   Button "Button_70" at 788,457 size 126x262; TextOff 'Text'
      on Release: function_efd93a16("Tank 2S Status", 168, 315, -1, 0, 1)
      Appearance <- "504_Tank Grouping_DB2020_RUN TANK 5"
   Button "Button_66" at 921,457 size 126x261; TextOff 'Text'
      on Release: function_efd93a16("Tank 1S Status", 168, 315, -1, 0, 1)
      Appearance <- "504_Tank Grouping_DB2020_RUN TANK 3"
   Button "Button_61" at 1093,328 size 130x248; TextOff 'Text'
      on Release: function_efd93a16("Tank FP Status", 168, 315, -1, 0, 1)
      Appearance <- "504_Tank Grouping_DB2020_RUN TANK 1"
   Button "Button_62" at 919,205 size 126x242; TextOff 'Text'
      on Release: function_efd93a16("Tank 1P Status", 168, 315, -1, 0, 1)
      Appearance <- "504_Tank Grouping_DB2020_RUN TANK 2"
   Button "Button_68" at 789,202 size 126x246; TextOff 'Text'
      on Release: function_efd93a16("Tank 2P Status", 168, 315, -1, 0, 1)
      Appearance <- "504_Tank Grouping_DB2020_RUN TANK 4"
   Button "Button_72" at 654,205 size 126x242; TextOff 'Text'
      on Release: function_efd93a16("Tank 3P Status", 168, 315, -1, 0, 1)
      Appearance <- "504_Tank Grouping_DB2020_RUN TANK 6"
   Button "Button_76" at 524,205 size 126x243; TextOff 'Text'
      on Release: function_efd93a16("Tank 4P Status", 168, 315, -1, 0, 1)
      Appearance <- "504_Tank Grouping_DB2020_RUN TANK 8"
   Button "Button_78" at 392,206 size 126x241; TextOff 'Text'
      on Release: function_efd93a16("Tank 5P Status", 168, 315, -1, 0, 1)
      Appearance <- "504_Tank Grouping_DB2020_RUN TANK 10"
   Button "Button_84" at 259,204 size 126x244; TextOff 'Text'
      on Release: function_efd93a16("Tank 6P Status", 168, 315, -1, 0, 1)
      Appearance <- "504_Tank Grouping_DB2020_RUN TANK 12"
   Group "Group_1" at 711,46 size 50x27; FormatPattern 999; Unit h
   Group "Group_2" at 605,46 size 57x27; FormatPattern 999; Unit h
   Button "HmiScreenItemData_5" at 180,144 size 116x50; TextOn 'Back'; TextOff 'Tank Status'
      on Release: function_efd93a16("Tank Status", 400, 250, -1, -1, 1)
   Button "Button_10" at 14,93 size 153x55; TextOff 'Text'
      on Release: function_efd93a16("Salinity - Acceptance", 168, 315, -1, 0, 1)
      Visibility <- "2068_Sys_Status_Data_SAL_VALID"
   Button "Button_12" at 14,93 size 153x54; TextOff 'Text'
      on Release: function_efd93a16("Tank Times", 300, 200, -1, 0, 1)
      Visibility <- "2068_Sys_Status_Data_Times Visibil"
   IOField "I/O field_29" at 664,46 size 45x27; FormatPattern 99; Unit h
      Visibility <- "2110_BTCS_CNTRL_DB_BTCS_STATE"
      ProcessValue <- "Sequence Times_DB_Treatment Timer_Hours Left"
   IOField "I/O field_30" at 664,46 size 45x27; FormatPattern 99; Unit h
      Visibility <- "2110_BTCS_CNTRL_DB_BTCS_STATE"
      ProcessValue <- "Sequence Times_DB_Pre-Dwell Timer_Hours Left"
   Button "Button_59" at 298,44 size 240x30; TextOn 'TB3 Enabled'; TextOff 'BWT System Shutting Down'
      Visibility <- "2110_BTCS_CNTRL_DB_BTCS_STATE"
   Button "Button_60" at 299,44 size 240x30; TextOn 'TB3 Enabled'; TextOff 'BWT System Enabled'
      Visibility <- "2110_BTCS_CNTRL_DB_BTCS_STATE"
   IOField "I/O field_15" at 711,46 size 50x27; FormatPattern 99; Unit m
      Visibility <- "2110_BTCS_CNTRL_DB_BTCS_STATE"
      ProcessValue <- "Sequence Times_DB_Treatment Timer_Minutes Left"
   IOField "I/O field_16" at 711,46 size 50x27; FormatPattern 99; Unit m
      Visibility <- "2110_BTCS_CNTRL_DB_BTCS_STATE"
      ProcessValue <- "Sequence Times_DB_Pre-Dwell Timer_Minutes Left"
   IOField "I/O field_17" at 605,46 size 57x27; FormatPattern 999; Unit d
      Visibility <- "2110_BTCS_CNTRL_DB_BTCS_STATE"
      ProcessValue <- "Sequence Times_DB_Treatment Timer_Days Left"
   IOField "I/O field_18" at 605,46 size 57x27; FormatPattern 999; Unit d
      Visibility <- "2110_BTCS_CNTRL_DB_BTCS_STATE"
      ProcessValue <- "Sequence Times_DB_Pre-Dwell Timer_Days Left"

screen "Balast Water Treatment Setup" 1280x800, template "Template"
   Button "HmiScreenItemData_1" at 1,1 size 150x40; TextOn 'Back'; TextOff 'Main Index'
      on Release: ActivateScreen("02 Main Index", 0)
   Button "HmiScreenItemData_8" at 276,83 size 219x27; TextOn 'Back'; TextOff 'Plant Operation'
   Button "HmiScreenItemData_23" at 282,116 size 150x47; TextOn 'Back'; TextOff 'Accept & Launch'; Authorization "Operate"
      Appearance <- "2110_BTCS_CNTRL_DB_BTCS_STATE"
      on Release: function_efd93a16("BWTS Start Confirm", 400, 200, -1, -1, 1)
      ObjectEnable <- "82_To_HMI_CRNT_MODE_GCU"
   Button "HmiScreenItemData_14" at 828,54 size 416x27; TextOn 'Back'; TextOff 'Treatment Durations'
   TextField "Text field_1" at 925,535 size 220x18; Text 'Tank Water Low Level (LT421)'
   TextField "Text field_2" at 925,573 size 220x18; Text 'Tank Water Low Level (LT422)'
   TextField "Text field_3" at 925,501 size 85x18; Text 'Description'
   TextField "Text field_5" at 925,611 size 215x18; Text 'De-Oxygenation DO Set Point'
   TextField "Text field_6" at 1164,501 size 67x18; Text 'Setpoint'
   Button "HmiScreenItemData_15" at 915,461 size 329x27; TextOn 'Back'; TextOff 'Ballast Tank Treatment Settings'
   IOField "I/O field_4" at 1153,530 size 80x28; Authorization "Operate"; FormatPattern 999.9; Unit  %
      ProcessValue <- "2084_Setpoints_LT421_Lo"
   IOField "I/O field_5" at 1153,568 size 80x28; Authorization "Operate"; FormatPattern 999.9; Unit  %
      ProcessValue <- "2084_Setpoints_LT422_Lo"
   IOField "I/O field_6" at 1153,606 size 80x28; Authorization "Operate"; FormatPattern 99.9; Unit  mg/l
      ProcessValue <- "2084_Setpoints_DO_SP"
   Button "HmiScreenItemData_16" at 482,461 size 334x27; TextOn 'Back'; TextOff 'Manual Ballast Tank Selection'
   Button "HmiScreenItemData_34" at 43,83 size 230x27; TextOn 'Back'; TextOff 'Plant Mode of Operation'
   Button "HmiScreenItemData_18" at 43,54 size 452x27; TextOn 'Back'; TextOff 'Ballast Water Treatment'
   Button "HmiScreenItemData_40" at 508,54 size 300x27; TextOn 'Back'; TextOff 'Treatment Status'
   TextField "Text field_14" at 837,94 size 85x18; Text 'Description'
   TextField "Text field_17" at 1054,94 size 67x18; Text 'Setpoint'
   IOField "I/O field_10" at 1040,132 size 92x27; Authorization "Operating Mode"; FormatPattern 999.99; Unit  Days
      ProcessValue <- "2115_VOYAGE_TIME_DAYS_VOYAGE_DAYS"
   IOField "I/O field_12" at 1040,267 size 79x28; Authorization "Commissioning"; FormatPattern 999; Unit  Hrs
      ProcessValue <- "2110_BTCS_CNTRL_DB_DE_OX_HRS"
   IOField "I/O field_13" at 1040,335 size 79x28; Authorization "Commissioning"; FormatPattern 999; Unit  Hrs
      ProcessValue <- "2110_BTCS_CNTRL_DB_DWELL_HRS"
   IOField "I/O field_14" at 1040,369 size 79x28; Authorization "Commissioning"; FormatPattern 999; Unit  Hrs
      ProcessValue <- "2110_BTCS_CNTRL_DB_RE_OX_HRS"
   IOField "I/O field_15" at 1040,403 size 79x28; Authorization "Commissioning"; FormatPattern 999; Unit  Hrs
      ProcessValue <- "2110_BTCS_CNTRL_DB_POST_DWELL_HRS"
   Button "HmiScreenItemData_11" at 836,128 size 203x35; TextOn 'Back'; TextOff 'Voyage A'
   Button "HmiScreenItemData_12" at 836,233 size 203x28; TextOn 'Back'; TextOff 'Pre Dwell Time'
   Button "HmiScreenItemData_13" at 836,267 size 203x28; TextOn 'Back'; TextOff 'De-Oxygenation Minimum Time'
   Button "HmiScreenItemData_43" at 836,335 size 203x28; TextOn 'Back'; TextOff 'Dwell Time'
   Button "HmiScreenItemData_44" at 836,369 size 203x28; TextOn 'Back'; TextOff 'Re-Oxygenation Time'
   Button "HmiScreenItemData_45" at 836,403 size 203x28; TextOn 'Back'; TextOff 'Post Dwell Time'
   IOField "I/O field_17" at 1060,169 size 79x28; Authorization "User administration"; FormatPattern 999; Unit  Hrs
      ProcessValue <- "2110_BTCS_CNTRL_DB_TOT_SEQ_HRS"
   Button "HmiScreenItemData_42" at 836,169 size 203x28; TextOn 'Back'; TextOff 'Total Treatment Time'
   Button "HmiScreenItemData_47" at 482,461 size 418x27; TextOn 'Back'; TextOff 'Automatic Ballast Tank Selection'
   Button "HmiScreenItemData_9" at 525,88 size 220x30; TextOn 'Back'; TextOff 'Pre Dwell Time Completed'
   Button "HmiScreenItemData_17" at 525,148 size 220x30; TextOn 'Back'; TextOff 'De-Oxygenation Completed'
   Button "HmiScreenItemData_38" at 525,178 size 220x30; TextOn 'Back'; TextOff 'Dwell Time Completed'
   Button "HmiScreenItemData_39" at 525,238 size 220x30; TextOn 'Back'; TextOff 'Re-Oxygenation Completed'
   Button "HmiScreenItemData_41" at 525,269 size 220x30; TextOn 'Back'; TextOff 'Post Dwell Time Completed'
   Button "HmiScreenItemData_46" at 525,118 size 220x30; TextOn 'Back'; TextOff 'Inert Gas Transfer Active'
   Button "HmiScreenItemData_48" at 525,208 size 220x30; TextOn 'Back'; TextOff 'Ambient Air Transfer Active'
   Button "HmiScreenItemData_52" at 525,118 size 220x30; TextOn 'Back'; TextOff 'IG Transfer Completed'
   Button "HmiScreenItemData_53" at 525,208 size 220x30; TextOn 'Back'; TextOff 'Ambient Air Transfer Completed'
   Button "HmiScreenItemData_3" at 1129,1 size 150x40; TextOn 'I&A Compressor Ok'; TextOff 'Back'
      on Release: function_efd93a16()
   TextField "Text field_11" at 1179,94 size 36x18; Text 'ETA'
   IOField "I/O field_16" at 1156,233 size 83x28; Authorization "User administration"; FormatPattern 999; Unit  min
      ProcessValue <- "2102_TIME_CALCS_DB_PRE_DWELL_MINS_RMNG"
   IOField "I/O field_18" at 1156,267 size 83x28; Authorization "User administration"; FormatPattern 999; Unit  min
   IOField "I/O field_19" at 1156,335 size 83x28; FormatPattern 999; Unit  min
      ProcessValue <- "2102_TIME_CALCS_DB_DWELL_MINS_RMNG"
   IOField "I/O field_20" at 1156,369 size 83x28; FormatPattern 999; Unit  min
      ProcessValue <- "2102_TIME_CALCS_DB_RE_OX_MINS_RMNG"
   IOField "I/O field_21" at 1156,403 size 83x28; FormatPattern 999; Unit  min
      ProcessValue <- "2102_TIME_CALCS_DB_POST_DWELL_MINS_RMNG"
   IOField "I/O field_22" at 1156,169 size 83x28; Authorization "User administration"; FormatPattern 999; Unit  Hrs
      ProcessValue <- "2110_BTCS_CNTRL_DB_RMNG_SEQ_HRS"
   Rectangle "Rectangle_25" at 281,165 size 179x59
      Visibility <- "2100_AUTO_SEQ_DB_SEQ_RNG"
   Button "HmiScreenItemData_4" at 282,172 size 150x47; TextOn 'Back'; TextOff 'Abort & Stop'; Authorization "Operate"
      Appearance <- "2110_BTCS_CNTRL_DB_BTCS_STATE"
      on Release: function_efd93a16("BWTS Stop Confirm", 400, 200, -1, -1, 1)
      ObjectEnable <- "82_To_HMI_CRNT_MODE_GCU"
   Circle "Circle_9" at 453,125 size 29x29
      Appearance <- "2110_BTCS_CNTRL_DB_BTCS_STATE"
   Circle "Circle_1" at 453,181 size 29x29
      Appearance <- "2110_BTCS_CNTRL_DB_BTCS_STATE"
   TextField "Text field_60" at 936,698 size 290x35; Text 'SALINITY ACCEPTED'
      Visibility <- "2068_Sys_Status_Data_SAL_VALID"
   Circle "Circle_19" at 220,233 size 29x29
      Appearance <- "150_GCU_LCL_CNTRL_DB_LCL_CNTRL_ACTV"
   Circle "Circle_20" at 220,180 size 29x29
      Appearance <- "82_To_HMI_CRNT_MODE_GCU"
   Button "HmiScreenItemData_36" at 49,170 size 150x51; TextOn 'Back'; TextOff 'Manual'; Authorization "Operate"
      on Press: function_b14e0dd5("80_From_HMI_Request_Manual", 0); ResetBit("150_GCU_LCL_CNTRL_DB_LCL_CNTRL_ACTV")
   Circle "Circle_21" at 220,126 size 29x29
      Appearance <- "82_To_HMI_CRNT_MODE_GCU"
   Button "HmiScreenItemData_37" at 49,116 size 150x51; TextOn 'Back'; TextOff 'Full Auto'; Authorization "Operate"
      on Press: function_b14e0dd5("80_From_HMI_Request_Auto", 0); ResetBit("150_GCU_LCL_CNTRL_DB_LCL_CNTRL_ACTV")
   Button "HmiScreenItemData_49" at 49,225 size 150x51; TextOn 'Back'; TextOff 'Local Auto'; Authorization "User administration"
      on Press: InvertBit("150_GCU_LCL_CNTRL_DB_LCL_CNTRL_ACTV"); function_b14e0dd5("80_From_HMI_Request_Auto", 0); ResetBit("80_From_HMI_Request_Manual")
   Circle "Circle_22" at 220,126 size 29x29
      Visibility <- "150_GCU_LCL_CNTRL_DB_LCL_CNTRL_ACTV"
   Circle "Circle_30" at 220,233 size 29x29
      Visibility <- "82_To_HMI_CRNT_MODE_GCU"
   Button "Button_4" at 493,507 size 100x23; TextOff 'FPT'; Authorization "Operate"
      on Press: function_b14e0dd5("504_Tank Grouping_DB2020_TANK ACTIV 1", 0)
      Appearance <- "504_Tank Grouping_DB2020_TANK ACTIV 1"
   Button "HmiScreenItemData_50" at 1156,297 size 83x35; TextOn 'Back'; TextOff 'Boost'; Authorization "Commissioning"
      on Press: InvertBit("Sequence Times_DB_Boost")
      Visibility <- "user_group"
      Appearance <- "Sequence Times_DB_Boost"
   IOField "I/O field_1" at 1040,301 size 79x28; Authorization "Commissioning"; FormatPattern 999; Unit  Hrs
      ProcessValue <- "2110_BTCS_CNTRL_DB_DE_OX_SP_HRS"
   Button "HmiScreenItemData_6" at 836,301 size 203x28; TextOn 'Back'; TextOff 'De-Oxygenation Setpoint Time'
   Rectangle "Rectangle_21" at 917,659 size 327x40
      Appearance <- "2068_Sys_Status_Data_SAL_VALID"
   TextField "Text field_48" at 916,664 size 128x30; Text 'Salinity Value:'
   IOField "I/O field_31" at 1036,664 size 74x30; FormatPattern 99.9; Unit psu
      ProcessValue <- "80_From_HMI_SAL_VALUE"
   Button "HmiScreenItemData_35" at 1108,664 size 135x30; TextOn 'Back'; TextOff 'Confirm Salinity'
      on Release: function_efd93a16("Salinity - Acceptance", 0, 0, 1, 3, 1)
   Group "Group_18" at 921,659 size 322x40
   Group "Group" at 916,659 size 327x40; Authorization "Operate"
   Button "HmiScreenItemData_7" at 1156,85 size 83x35; TextOn 'CONTINUE'; TextOff 'Continue'; Authorization "Operating Mode"
      on Press: InvertBit("80_From_HMI_TIMER RST Supres")
      Appearance <- "80_From_HMI_TIMER RST Supres"
   IOField "I/O field_25" at 1040,201 size 79x28; Authorization "User administration"; FormatPattern 999.9; Unit  Hrs
      ProcessValue <- "504_Tank Grouping_DB2020_Sequence Time m Offset_Real"
   Button "HmiScreenItemData_2" at 836,201 size 203x28; TextOn 'Back'; TextOff 'Differential Treatment Time'
   IOField "I/O field_3" at 1156,201 size 83x28; Authorization "User administration"; FormatPattern 999; Unit  min
      ProcessValue <- "504_Tank Grouping_DB2020_Diff Time Remain"
   Button "Button_1" at 817,594 size 79x32; TextOff '3'; Authorization "Operate"
      on Press: function_b14e0dd5("504_Tank Grouping_DB2020_GROUP ACTIV 3", 0)
      Appearance <- "504_Tank Grouping_DB2020_GROUP ACTIVE INT 3"
   Button "Button_2" at 817,628 size 79x32; TextOff '4'; Authorization "Operate"
      on Press: function_b14e0dd5("504_Tank Grouping_DB2020_GROUP ACTIV 4", 0)
      Appearance <- "504_Tank Grouping_DB2020_GROUP ACTIVE INT 4"
   Button "Button_10" at 818,662 size 79x32; TextOff '5'; Authorization "Operate"
      on Press: function_b14e0dd5("504_Tank Grouping_DB2020_GROUP ACTIV 5", 0)
      Appearance <- "504_Tank Grouping_DB2020_GROUP ACTIVE INT 5"
   Button "Button_11" at 818,696 size 79x32; TextOff '6'; Authorization "Operate"
      on Press: function_b14e0dd5("504_Tank Grouping_DB2020_GROUP ACTIV 6", 0)
      Appearance <- "504_Tank Grouping_DB2020_GROUP ACTIVE INT 6"
   Button "Button_12" at 818,731 size 79x32; TextOff '7'; Authorization "Operate"
      on Press: function_b14e0dd5("504_Tank Grouping_DB2020_GROUP ACTIV 7", 0)
      Appearance <- "504_Tank Grouping_DB2020_GROUP ACTIVE INT 7"
   IOField "I/O field_37" at 183,323 size 90x29; Authorization "Commissioning"; FormatPattern 999; Unit  step
      ProcessValue <- "2110_BTCS_CNTRL_DB_BTCS_STEP"
   Button "HmiScreenItemData_10" at 43,323 size 137x29; TextOn 'Back'; TextOff 'BWTS Step'
   Button "HmiScreenItemData_51" at 43,358 size 137x29; TextOn 'Back'; TextOff 'BWTS State'
   Button "HmiScreenItemData_54" at 276,323 size 532x29; TextOn 'Back'; TextOff 'IGG STEP'; TextList "STEP LIST BTCS"
      ProcessValue <- "2110_BTCS_CNTRL_DB_BTCS_STEP"
   Button "HmiScreenItemData_55" at 276,358 size 532x29; TextOn 'Back'; TextOff 'IGG STEP'; TextList "STATE LIST BTCS"
      ProcessValue <- "2110_BTCS_CNTRL_DB_BTCS_STATE"
   Circle "Circle_2" at 421,496 size 26x26
      Appearance <- "80_From_HMI_BWT_BYPASS"
   Button "HmiScreenItemData_57" at 88,494 size 304x33; TextOn 'Back'; TextOff 'Ballast Water Treatment'; Authorization "Operate"
      on Press: InvertBit("80_From_HMI_BWT_BYPASS(1)"); ResetBit("80_From_HMI_CRG_BLNK_MODE(1)")
      Appearance <- "80_From_HMI_BWT_BYPASS(1)"
      ObjectEnable <- "100_GCU_AUTO_SEQ_DB_CRNT_STEP"
   Circle "Circle_3" at 421,534 size 26x26
      Appearance <- "80_From_HMI_CRG_BLNK_MODE"
   Button "HmiScreenItemData_58" at 88,532 size 304x33; TextOn 'Back'; TextOff 'Cargo Blanketing'; Authorization "Operate"
      on Press: InvertBit("80_From_HMI_CRG_BLNK_MODE(1)"); ResetBit("80_From_HMI_BWT_BYPASS(1)")
      Appearance <- "80_From_HMI_CRG_BLNK_MODE(1)"
      ObjectEnable <- "100_GCU_AUTO_SEQ_DB_CRNT_STEP"
   Button "HmiScreenItemData_56" at 41,461 size 425x27; TextOn 'Back'; TextOff 'Inert Gas Transfer Mode'
   Button "Button_7" at 817,526 size 79x32; TextOff '1'; Authorization "Operate"
      on Press: function_b14e0dd5("504_Tank Grouping_DB2020_GROUP ACTIV 1", 0)
      Appearance <- "504_Tank Grouping_DB2020_GROUP ACTIVE INT 1"
   Button "Button_8" at 817,560 size 79x32; TextOff '2'; Authorization "Operate"
      on Press: function_b14e0dd5("504_Tank Grouping_DB2020_GROUP ACTIV 2", 0)
      Appearance <- "504_Tank Grouping_DB2020_GROUP ACTIVE INT 2"
   Button "Button_9" at 493,539 size 100x23; TextOff 'TANK - 1P'; Authorization "Operate"
      on Press: function_b14e0dd5("504_Tank Grouping_DB2020_TANK ACTIV 2", 0)
      Appearance <- "504_Tank Grouping_DB2020_TANK ACTIV 2"
   Button "Button_14" at 493,571 size 100x23; TextOff 'TANK - 2P'; Authorization "Operate"
      on Press: function_b14e0dd5("504_Tank Grouping_DB2020_TANK ACTIV 4", 0)
      Appearance <- "504_Tank Grouping_DB2020_TANK ACTIV 4"
   Button "Button_15" at 493,603 size 100x23; TextOff 'TANK - 3P'; Authorization "Operate"
      on Press: function_b14e0dd5("504_Tank Grouping_DB2020_TANK ACTIV 6", 0)
      Appearance <- "504_Tank Grouping_DB2020_TANK ACTIV 6"
   Button "Button_16" at 493,636 size 100x23; TextOff 'TANK - 4P'; Authorization "Operate"
      on Press: function_b14e0dd5("504_Tank Grouping_DB2020_TANK ACTIV 8", 0)
      Appearance <- "504_Tank Grouping_DB2020_TANK ACTIV 8"
   Button "Button_17" at 493,668 size 100x23; TextOff 'TANK - 5P'; Authorization "Operate"
      on Press: function_b14e0dd5("504_Tank Grouping_DB2020_TANK ACTIV 10", 0)
      Appearance <- "504_Tank Grouping_DB2020_TANK ACTIV 10"
   Button "Button_18" at 493,700 size 100x23; TextOff 'TANK - 6P'; Authorization "Operate"
      on Press: function_b14e0dd5("504_Tank Grouping_DB2020_TANK ACTIV 12", 0)
      Appearance <- "504_Tank Grouping_DB2020_TANK ACTIV 12"
   Button "Button_19" at 493,733 size 100x23; TextOff 'TANK - APT'; Authorization "Operate"
      on Press: function_b14e0dd5("504_Tank Grouping_DB2020_TANK ACTIV 14", 0)
      Appearance <- "504_Tank Grouping_DB2020_TANK ACTIV 14"
   Button "Button_20" at 706,539 size 100x23; TextOff 'TANK - 1S'; Authorization "Operate"
      on Press: function_b14e0dd5("504_Tank Grouping_DB2020_TANK ACTIV 3", 0)
      Appearance <- "504_Tank Grouping_DB2020_TANK ACTIV 3"
   Button "Button_21" at 706,571 size 100x23; TextOff 'TANK - 2S'; Authorization "Operate"
      on Press: function_b14e0dd5("504_Tank Grouping_DB2020_TANK ACTIV 5", 0)
      Appearance <- "504_Tank Grouping_DB2020_TANK ACTIV 5"
   Button "Button_22" at 706,603 size 100x23; TextOff 'TANK - 3S'; Authorization "Operate"
      on Press: function_b14e0dd5("504_Tank Grouping_DB2020_TANK ACTIV 7", 0)
      Appearance <- "504_Tank Grouping_DB2020_TANK ACTIV 7"
   Button "Button_23" at 706,635 size 100x23; TextOff 'TANK - 4S'; Authorization "Operate"
      on Press: function_b14e0dd5("504_Tank Grouping_DB2020_TANK ACTIV 9", 0)
      Appearance <- "504_Tank Grouping_DB2020_TANK ACTIV 9"
   Button "Button_24" at 706,667 size 100x23; TextOff 'TANK - 5S'; Authorization "Operate"
      on Press: function_b14e0dd5("504_Tank Grouping_DB2020_TANK ACTIV 11", 0)
      Appearance <- "504_Tank Grouping_DB2020_TANK ACTIV 11"
   Button "Button_25" at 706,700 size 100x23; TextOff 'TANK - 6S'; Authorization "Operate"
      on Press: function_b14e0dd5("504_Tank Grouping_DB2020_TANK ACTIV 13", 0)
      Appearance <- "504_Tank Grouping_DB2020_TANK ACTIV 13"
   IOField "I/O field_38" at 183,358 size 90x29; Authorization "Commissioning"; FormatPattern 9; Unit  state
      ProcessValue <- "2110_BTCS_CNTRL_DB_BTCS_STATE"
   Switch "Switch_8" at 776,732 size 32x29; CaptionText 'Switch'; TextOn 'ON'; TextOff 'OFF'; Authorization "User administration"; PictureOff "Design_5_PilotLight_Green_Off"; PictureOn "Design_5_PilotLight_Green_On"
      on Change: InvertBit("80_From_HMI_Test Tank Request")
      ProcessValue <- "504_Tank Grouping_DB2020_RUN"
      Visibility <- "user_group"
   Circle "Circle_31" at 621,507 size 20x20
      Visibility <- "504_Tank Grouping_DB2020_RUN TANK 1"
      Appearance <- "504_Tank Grouping_DB2020_RUN TANK 1"
   Circle "Circle_4" at 600,573 size 20x20
      Appearance <- "504_Tank Grouping_DB2020_GROUP of TANK 4"
   Circle "Circle_6" at 599,604 size 20x20
      Appearance <- "504_Tank Grouping_DB2020_GROUP of TANK 6"
   Circle "Circle_7" at 599,541 size 20x20
      Appearance <- "504_Tank Grouping_DB2020_GROUP of TANK 2"
   Circle "Circle_8" at 599,669 size 20x20
      Appearance <- "504_Tank Grouping_DB2020_GROUP of TANK 10"
   Circle "Circle_10" at 599,637 size 20x20
      Appearance <- "504_Tank Grouping_DB2020_GROUP of TANK 8"
   Circle "Circle_11" at 599,734 size 20x20
      Appearance <- "504_Tank Grouping_DB2020_GROUP of TANK 14"
   Circle "Circle_12" at 599,701 size 20x20
      Appearance <- "504_Tank Grouping_DB2020_GROUP of TANK 12"
   IOField "I/O field_8" at 599,544 size 20x14; FormatPattern 99
      ProcessValue <- "504_Tank Grouping_DB2020_GROUP of TANK 2"
   IOField "I/O field_9" at 599,576 size 20x14; FormatPattern 99
      ProcessValue <- "504_Tank Grouping_DB2020_GROUP of TANK 4"
   IOField "I/O field_26" at 599,607 size 20x14; FormatPattern 99
      ProcessValue <- "504_Tank Grouping_DB2020_GROUP of TANK 6"
   IOField "I/O field_28" at 599,640 size 20x14; FormatPattern 99
      ProcessValue <- "504_Tank Grouping_DB2020_GROUP of TANK 8"
   IOField "I/O field_30" at 599,672 size 20x14; FormatPattern 99
      ProcessValue <- "504_Tank Grouping_DB2020_GROUP of TANK 10"
   IOField "I/O field_33" at 599,704 size 20x14; FormatPattern 99
      ProcessValue <- "504_Tank Grouping_DB2020_GROUP of TANK 12"
   IOField "I/O field_35" at 599,737 size 20x14; FormatPattern 99
      ProcessValue <- "504_Tank Grouping_DB2020_GROUP of TANK 14"
   Circle "Circle_13" at 678,573 size 20x20
      Appearance <- "504_Tank Grouping_DB2020_GROUP of TANK 5"
   Circle "Circle_14" at 678,603 size 20x20
      Appearance <- "504_Tank Grouping_DB2020_GROUP of TANK 7"
   Circle "Circle_15" at 678,541 size 20x20
      Appearance <- "504_Tank Grouping_DB2020_GROUP of TANK 3"
   Circle "Circle_16" at 678,668 size 20x20
      Appearance <- "504_Tank Grouping_DB2020_GROUP of TANK 11"
   Circle "Circle_17" at 678,636 size 20x20
      Appearance <- "504_Tank Grouping_DB2020_GROUP of TANK 9"
   Circle "Circle_18" at 678,701 size 20x20
      Appearance <- "504_Tank Grouping_DB2020_GROUP of TANK 13"
   IOField "I/O field_23" at 678,544 size 20x14; FormatPattern 99
      ProcessValue <- "504_Tank Grouping_DB2020_GROUP of TANK 3"
   IOField "I/O field_24" at 678,576 size 20x14; FormatPattern 99
      ProcessValue <- "504_Tank Grouping_DB2020_GROUP of TANK 5"
   IOField "I/O field_27" at 678,606 size 20x14; FormatPattern 99
      ProcessValue <- "504_Tank Grouping_DB2020_GROUP of TANK 7"
   IOField "I/O field_29" at 678,639 size 20x14; FormatPattern 99
      ProcessValue <- "504_Tank Grouping_DB2020_GROUP of TANK 9"
   IOField "I/O field_32" at 678,671 size 20x14; FormatPattern 99
      ProcessValue <- "504_Tank Grouping_DB2020_GROUP of TANK 11"
   IOField "I/O field_34" at 678,704 size 20x14; FormatPattern 99
      ProcessValue <- "504_Tank Grouping_DB2020_GROUP of TANK 13"
   Circle "Circle_32" at 621,540 size 20x20
      Visibility <- "504_Tank Grouping_DB2020_RUN TANK 2"
      Appearance <- "504_Tank Grouping_DB2020_RUN TANK 2"
   Circle "Circle_33" at 656,540 size 20x20
      Visibility <- "504_Tank Grouping_DB2020_RUN TANK 3"
      Appearance <- "504_Tank Grouping_DB2020_RUN TANK 3"
   Circle "Circle_34" at 621,572 size 20x20
      Visibility <- "504_Tank Grouping_DB2020_RUN TANK 4"
      Appearance <- "504_Tank Grouping_DB2020_RUN TANK 4"
   Circle "Circle_35" at 656,572 size 20x20
      Visibility <- "504_Tank Grouping_DB2020_RUN TANK 5"
      Appearance <- "504_Tank Grouping_DB2020_RUN TANK 5"
   Circle "Circle_36" at 621,604 size 20x20
      Visibility <- "504_Tank Grouping_DB2020_RUN TANK 6"
      Appearance <- "504_Tank Grouping_DB2020_RUN TANK 6"
   Circle "Circle_37" at 656,604 size 20x20
      Visibility <- "504_Tank Grouping_DB2020_RUN TANK 7"
      Appearance <- "504_Tank Grouping_DB2020_RUN TANK 7"
   Circle "Circle_38" at 621,636 size 20x20
      Visibility <- "504_Tank Grouping_DB2020_RUN TANK 8"
      Appearance <- "504_Tank Grouping_DB2020_RUN TANK 8"
   Circle "Circle_39" at 656,636 size 20x20
      Visibility <- "504_Tank Grouping_DB2020_RUN TANK 9"
      Appearance <- "504_Tank Grouping_DB2020_RUN TANK 9"
   Circle "Circle_40" at 621,668 size 20x20
      Visibility <- "504_Tank Grouping_DB2020_RUN TANK 10"
      Appearance <- "504_Tank Grouping_DB2020_RUN TANK 10"
   Circle "Circle_41" at 656,668 size 20x20
      Visibility <- "504_Tank Grouping_DB2020_RUN TANK 11"
      Appearance <- "504_Tank Grouping_DB2020_RUN TANK 11"
   Circle "Circle_42" at 621,701 size 20x20
      Visibility <- "504_Tank Grouping_DB2020_RUN TANK 12"
      Appearance <- "504_Tank Grouping_DB2020_RUN TANK 12"
   Circle "Circle_43" at 656,701 size 20x20
      Visibility <- "504_Tank Grouping_DB2020_RUN TANK 13"
      Appearance <- "504_Tank Grouping_DB2020_RUN TANK 13"
   Circle "Circle_44" at 621,733 size 20x20
      Visibility <- "504_Tank Grouping_DB2020_RUN TANK 14"
      Appearance <- "504_Tank Grouping_DB2020_RUN TANK 14"
   TextField "Text field_7" at 648,740 size 136x18; Text 'Test Tank Request'
      Visibility <- "user_group"
   Rectangle "Rectangle_6" at 816,488 size 82x37
      Visibility <- "504_Tank Grouping_DB2020_SetGroupSR"
   Button "Button_13" at 819,491 size 76x31; TextOff 'Set Group'; Authorization "Parameter Change"
      on Press: function_b14e0dd5("504_Tank Grouping_DB2020_SetGroup", 0)
      Appearance <- "504_Tank Grouping_DB2020_GROUP SET"
   Button "HmiScreenItemData_5" at 41,576 size 426x27; TextOn 'Back'; TextOff 'Automatic Gas to Tank Valves Cycling'
   Button "HmiScreenItemData_19" at 370,722 size 83x35; TextOn 'ENABLE'; TextOff 'Enable'; Authorization "Operate"
      on Press: InvertBit("504_Tank Grouping_DB2020_Valve Cycle_Enable")
      Appearance <- "504_Tank Grouping_DB2020_Valve Cycle_Enable"
   TextField "Text field_8" at 54,652 size 254x18; Text 'Gas to Tank Valves Cycle Frequency'
   TextField "Text field_9" at 54,690 size 233x18; Text 'Gas to Tank Valves Cycle Length'
   TextField "Text field_10" at 54,618 size 85x18; Text 'Description'
   TextField "Text field_12" at 311,618 size 67x18; Text 'Setpoint'
   IOField "I/O field_39" at 310,649 size 70x28; Authorization "Operate"; FormatPattern 999; Unit h
      ProcessValue <- "504_Tank Grouping_DB2020_Valve Cycle_Period"
   IOField "I/O field_40" at 310,685 size 70x28; Authorization "Operate"; FormatPattern 9999; Unit s
      ProcessValue <- "504_Tank Grouping_DB2020_Valve Cycle_Length"
   TextField "Text field_13" at 385,618 size 58x18; Text 'Elapsed'
   IOField "I/O field_41" at 384,649 size 70x28; Authorization "Operate"; FormatPattern 999; Unit h
      ProcessValue <- "504_Tank Grouping_DB2020_Cycle Period_ET"
   IOField "I/O field_42" at 384,685 size 70x28; Authorization "Operate"; FormatPattern 9999; Unit s
      ProcessValue <- "504_Tank Grouping_DB2020_Cycle Length_ET"
   IOField "I/O field_48" at 1172,169 size 33x28; Authorization "User administration"; FormatPattern 99; Unit h
      ProcessValue <- "Sequence Times_DB_Treatment Timer_Hours Left"
   IOField "I/O field_51" at 1140,169 size 33x28; Authorization "User administration"; FormatPattern 99; Unit d
      ProcessValue <- "Sequence Times_DB_Treatment Timer_Days Left"
   IOField "I/O field_52" at 1204,169 size 35x28; Authorization "User administration"; FormatPattern 99; Unit m
      ProcessValue <- "Sequence Times_DB_Treatment Timer_Minutes Left"
   IOField "I/O field_43" at 1156,201 size 83x28; Authorization "User administration"; FormatPattern 999; Unit  min
      ProcessValue <- "504_Tank Grouping_DB2020_Diff Time Remain"
      Visibility <- "AlwaysTRUE"
   IOField "I/O field_44" at 1204,233 size 35x28; Authorization "User administration"; FormatPattern 99; Unit m
      ProcessValue <- "Sequence Times_DB_Pre-Dwell Timer_Minutes Left"
   IOField "I/O field_45" at 1172,233 size 33x28; Authorization "User administration"; FormatPattern 99; Unit h
      ProcessValue <- "Sequence Times_DB_Pre-Dwell Timer_Hours Left"
   IOField "I/O field_46" at 1140,233 size 33x28; Authorization "User administration"; FormatPattern 99; Unit d
      ProcessValue <- "Sequence Times_DB_Pre-Dwell Timer_Days Left"
   IOField "I/O field_47" at 1040,132 size 92x28; Authorization "Operating Mode"; FormatPattern 999.9; Unit  Days
      ProcessValue <- "Sequence Times_DB_Jurney Time"
   IOField "I/O field_49" at 1072,169 size 33x28; Authorization "User administration"; FormatPattern 99; Unit h
      ProcessValue <- "Sequence Times_DB_Treatment Timer_Hours"
   IOField "I/O field_50" at 1040,169 size 33x28; Authorization "User administration"; FormatPattern 99; Unit d
      ProcessValue <- "Sequence Times_DB_Treatment Timer_Days"
   IOField "I/O field_53" at 1104,169 size 35x28; Authorization "User administration"; FormatPattern 99; Unit m
      ProcessValue <- "Sequence Times_DB_Treatment Timer_Minutes"
   IOField "I/O field_54" at 1172,132 size 33x28; Authorization "User administration"; FormatPattern 99; Unit h
      ProcessValue <- "Sequence Times_DB_Jurney Timer_Hours Left"
   IOField "I/O field_55" at 1133,132 size 40x28; Authorization "User administration"; FormatPattern 999; Unit d
      ProcessValue <- "Sequence Times_DB_Jurney Timer_Days Left"
   IOField "I/O field_56" at 1204,132 size 35x28; Authorization "User administration"; FormatPattern 99; Unit m
      ProcessValue <- "Sequence Times_DB_Jurney Timer_Minutes Left"
   IOField "I/O field_57" at 1040,233 size 79x28; Authorization "Commissioning"; FormatPattern 9999.9; Unit  Hrs
      ProcessValue <- "Sequence Times_DB_Pre-Dwell Time"
   IOField "I/O field_58" at 1040,267 size 79x28; Authorization "Commissioning"; FormatPattern 999.9; Unit  Hrs
      ProcessValue <- "Sequence Times_DB_De-Ox Time"
   IOField "I/O field_59" at 1204,267 size 35x28; Authorization "User administration"; FormatPattern 99; Unit m
      ProcessValue <- "Sequence Times_DB_De-Ox Timer_Minutes Left"
   IOField "I/O field_60" at 1172,267 size 33x28; Authorization "User administration"; FormatPattern 99; Unit h
      ProcessValue <- "Sequence Times_DB_De-Ox Timer_Hours Left"
   IOField "I/O field_61" at 1140,267 size 33x28; Authorization "User administration"; FormatPattern 99; Unit d
      ProcessValue <- "Sequence Times_DB_De-Ox Timer_Days Left"
   IOField "I/O field_62" at 1040,301 size 79x28; Authorization "Commissioning"; FormatPattern 999.9; Unit  Hrs
      ProcessValue <- "Sequence Times_DB_De-Ox SP Time"
   IOField "I/O field_63" at 1040,335 size 79x28; Authorization "Commissioning"; FormatPattern 999.9; Unit  Hrs
      ProcessValue <- "Sequence Times_DB_Dwell Time"
   IOField "I/O field_64" at 1204,335 size 35x28; Authorization "User administration"; FormatPattern 99; Unit m
      ProcessValue <- "Sequence Times_DB_Dwell Timer_Minutes Left"
   IOField "I/O field_65" at 1172,335 size 33x28; Authorization "User administration"; FormatPattern 99; Unit h
      ProcessValue <- "Sequence Times_DB_Dwell Timer_Hours Left"
   IOField "I/O field_66" at 1140,335 size 33x28; Authorization "User administration"; FormatPattern 99; Unit d
      ProcessValue <- "Sequence Times_DB_Dwell Timer_Days Left"
   IOField "I/O field_2" at 1040,369 size 79x28; Authorization "Commissioning"; FormatPattern 999.9; Unit  Hrs
      ProcessValue <- "Sequence Times_DB_Re-Ox Time"
   IOField "I/O field_67" at 1204,369 size 35x28; Authorization "User administration"; FormatPattern 99; Unit m
      ProcessValue <- "Sequence Times_DB_Re-Ox Timer_Minutes Left"
   IOField "I/O field_68" at 1172,369 size 33x28; Authorization "User administration"; FormatPattern 99; Unit h
      ProcessValue <- "Sequence Times_DB_Re-Ox Timer_Hours Left"
   IOField "I/O field_69" at 1140,369 size 33x28; Authorization "User administration"; FormatPattern 99; Unit d
      ProcessValue <- "Sequence Times_DB_Re-Ox Timer_Days Left"
   IOField "I/O field_70" at 1040,403 size 79x28; Authorization "Commissioning"; FormatPattern 999.9; Unit  Hrs
      ProcessValue <- "Sequence Times_DB_Post-Dwell Time"
   IOField "I/O field_71" at 1204,403 size 35x28; Authorization "User administration"; FormatPattern 99; Unit m
      ProcessValue <- "Sequence Times_DB_Post-Dwell Timer_Minutes Left"
   IOField "I/O field_72" at 1172,403 size 33x28; Authorization "User administration"; FormatPattern 99; Unit h
      ProcessValue <- "Sequence Times_DB_Post-Dwell Timer_Hours Left"
   IOField "I/O field_73" at 1140,403 size 33x28; Authorization "User administration"; FormatPattern 99; Unit d
      ProcessValue <- "Sequence Times_DB_Post-Dwell Timer_Days Left"
   TextField "Text field_15" at 621,419 size 156x18; Text 'Treatment Timer Test'
      Visibility <- "user_group"
   Switch "Switch_1" at 774,411 size 32x29; CaptionText 'Switch'; TextOn 'ON'; TextOff 'OFF'; Authorization "User administration"; PictureOff "Design_5_PilotLight_Green_Off"; PictureOn "Design_5_PilotLight_Green_On"
      on Change: InvertBit("80_From_HMI_Jurney Start Simulator")
      Visibility <- "user_group"
      ProcessValue <- "80_From_HMI_Jurney Start Simulator"
   Circle "Circle_5" at 599,507 size 20x20
      Appearance <- "504_Tank Grouping_DB2020_GROUP of TANK 1"
   IOField "I/O field_7" at 599,510 size 20x14; FormatPattern 99
      ProcessValue <- "504_Tank Grouping_DB2020_GROUP of TANK 1"
   TextField "Text field_16" at 72,422 size 76x18; Text 'HeartBeat'
      Visibility <- "user_group"
   TextField "Text field_18" at 201,422 size 107x18; Text 'PLC HeartBeat'
      Visibility <- "user_group"
   Circle "Circle_45" at 40,414 size 26x26
      Appearance <- "CCR HMI HEART BEAT"
      Visibility <- "user_group"
   Circle "Circle_46" at 166,414 size 26x26
      Appearance <- "IGG PLC HEART BEAT"
      Visibility <- "user_group"
   TextField "Text field_19" at 445,403 size 133x18; Text 'Log IGG Simulator'
      Visibility <- "user_group"
   Switch "Switch_2" at 568,393 size 32x29; CaptionText 'Switch'; TextOn 'ON'; TextOff 'OFF'; Authorization "User administration"; PictureOff "Design_5_PilotLight_Green_Off"; PictureOn "Design_5_PilotLight_Green_On"
      on Change: InvertBit("68_Sys_Status_Data_LOG IGG Simulator")
      Visibility <- "user_group"
      ProcessValue <- "68_Sys_Status_Data_LOG IGG Simulator"
   TextField "Text field_20" at 445,435 size 136x18; Text 'Log GCU Simulator'
      Visibility <- "user_group"
   Switch "Switch_3" at 568,425 size 32x29; CaptionText 'Switch'; TextOn 'ON'; TextOff 'OFF'; Authorization "User administration"; PictureOff "Design_5_PilotLight_Green_Off"; PictureOn "Design_5_PilotLight_Green_On"
      on Change: InvertBit("68_Sys_Status_Data_LOG GCU Simulator")
      Visibility <- "user_group"
      ProcessValue <- "68_Sys_Status_Data_LOG GCU Simulator"
   Button "Button_5" at 53,722 size 210x35; TextOff 'PGC Setpoint Protection'
      on Press: function_efd93a16("PGC Setpoint Protection", 400, 200, -1, -1, 1)
   Button "Button_26" at 281,116 size 208x107; TextOff 'Text'
      on Release: function_efd93a16("Salinity - Acceptance", 168, 315, -1, 0, 1)
      Visibility <- "2068_Sys_Status_Data_SAL_VALID"
   Button "Button_27" at 280,115 size 204x107; TextOff 'Text'
      on Release: function_efd93a16("Tank Times", 300, 200, -1, 0, 1)
      Visibility <- "2068_Sys_Status_Data_Times Visibil"
   Group "Group_1" at 909,732 size 329x37
   IOField "I/O field_11" at 1156,201 size 83x28; Authorization "User administration"; FormatPattern 999; Unit  Hrs
      ProcessValue <- "2110_BTCS_CNTRL_DB_RMNG_SEQ_HRS"
   IOField "I/O field_74" at 1172,201 size 33x28; Authorization "User administration"; FormatPattern 99; Unit h
      ProcessValue <- "Sequence Times_DB_Offset Timer_Hours Left"
   IOField "I/O field_75" at 1140,201 size 33x28; Authorization "User administration"; FormatPattern 99; Unit d
      ProcessValue <- "Sequence Times_DB_Offset Timer_Days Left"
   IOField "I/O field_76" at 1204,201 size 35x28; Authorization "User administration"; FormatPattern 99; Unit m
      ProcessValue <- "Sequence Times_DB_Offset Timer_Minutes Left"
   Circle "Circle_23" at 764,91 size 24x24
      Appearance <- "2110_BTCS_CNTRL_DB_BTCS_STEP"
   Circle "Circle_24" at 764,120 size 24x24
      Appearance <- "100_GCU_AUTO_SEQ_DB_CRNT_STEP"
   Circle "Circle_25" at 764,150 size 24x24
      Appearance <- "2110_BTCS_CNTRL_DB_BTCS_STEP"
   Circle "Circle_26" at 764,180 size 24x24
      Appearance <- "2110_BTCS_CNTRL_DB_BTCS_STEP"
   Circle "Circle_27" at 764,210 size 24x24
      Appearance <- "100_GCU_AUTO_SEQ_DB_CRNT_STEP"
   Circle "Circle_28" at 764,240 size 24x24
      Appearance <- "2110_BTCS_CNTRL_DB_BTCS_STEP"
   Circle "Circle_29" at 764,270 size 24x24
      Appearance <- "2110_BTCS_CNTRL_DB_BTCS_STEP"
   TextField "Text field_34" at 980,733 size 187x35; Text 'TIMES VALID'
      Visibility <- "2102_TIME_CALCS_DB_TIMES_VALID"
   TextField "Text field_4" at 909,732 size 329x37; Text 'TIMES INVALID'
      Visibility <- "2102_TIME_CALCS_DB_TIMES_VALID"
   Rectangle "Rectangle_27" at 921,659 size 322x40
      Visibility <- "2068_Sys_Status_Data_SAL_CNF_CHK"
   TextField "Text field_62" at 925,664 size 156x30; Text 'Confirm Salinity? :'
      Visibility <- "2068_Sys_Status_Data_SAL_CNF_CHK"
   Button "Button_6" at 1086,664 size 67x30; TextOff 'YES'
      on Press: function_b14e0dd5("80_From_HMI_LOW_SAL_ACPT", 0)
      Visibility <- "2068_Sys_Status_Data_SAL_CNF_CHK"
   Button "Button_3" at 1166,664 size 67x30; TextOff 'NO'
      on Press: function_b14e0dd5("80_From_HMI_LOW_SAL_RJCT", 0)
      Visibility <- "2068_Sys_Status_Data_SAL_CNF_CHK"
   Rectangle "Rectangle_28" at 916,659 size 327x40
      Visibility <- "2100_AUTO_SEQ_DB_SEQ_RNG"
      Appearance <- "2102_TIME_CALCS_DB_RE_OX_SP_TMR_DN"
   TextField "Text field_49" at 920,664 size 211x30; Text 'Salinity Value :'
      Visibility <- "2100_AUTO_SEQ_DB_SEQ_RNG"
   IOField "I/O field_36" at 1131,664 size 95x30; Authorization "Operate"; FormatPattern 99.9; Unit psu
      ProcessValue <- "80_From_HMI_SAL_VALUE"
      Visibility <- "2100_AUTO_SEQ_DB_SEQ_RNG"

PopupScreen "Tank 1P Status" 885x425
   TrendView "Trend view_1" at 280,8 size 600x360
   TextField "Text field_4" at 20,136 size 86x22; Text 'Pressure:'
   IOField "I/O field_1" at 175,131 size 90x25; FormatPattern s999.9; Unit  mBar
      ProcessValue <- "20_TANKS_IP_DATA_RIO_01_FIRST_TANK_TANKS_PRESS"
   TextField "Text field_5" at 20,170 size 113x22; Text 'Water Level:'
   IOField "I/O field_2" at 175,165 size 90x25; FormatPattern 999.9; Unit  %
      ProcessValue <- "20_TANKS_IP_DATA_RIO_01_SECOND_TANK_BWT_LEVEL"
   TextField "Text field_6" at 20,204 size 137x22; Text 'MBG Flow Rate:'
   IOField "I/O field_3" at 175,199 size 90x25; FormatPattern 999.9; Unit  m³/hr
      ProcessValue <- "20_TANKS_IP_DATA_RIO_01_SECOND_TANK_MBG_FLOW"
   TextField "Text field_7" at 20,238 size 135x22; Text 'USD Flow Rate:'
   IOField "I/O field_4" at 175,233 size 90x25; FormatPattern 999.9; Unit  m³/hr
      ProcessValue <- "20_TANKS_IP_DATA_RIO_01_SECOND_TANK_USD_FLOW"
   TextField "Text field_8" at 20,272 size 140x22; Text 'Water pH Level:'
   IOField "I/O field_5" at 175,267 size 90x25; FormatPattern 99.9
      ProcessValue <- "20_TANKS_IP_DATA_RIO_01_SECOND_TANK_BWT_PH"
   TextField "Text field_9" at 20,306 size 143x22; Text 'Water DO Level:'
   IOField "I/O field_6" at 175,301 size 90x25; FormatPattern 99.99; Unit  mg/l
      ProcessValue <- "20_TANKS_IP_DATA_RIO_01_SECOND_TANK_BWT_DO"
   TextField "Text field_10" at 20,340 size 174x22; Text 'Water Temperature:'
   IOField "I/O field_7" at 190,335 size 75x25; FormatPattern 999.9; Unit  °C
      ProcessValue <- "20_TANKS_IP_DATA_RIO_01_SECOND_TANK_BWT_TEMP"
   Button "Button_1" at 51,5 size 219x35; TextOff 'Port Tank 1 (1P)'
      on Release: function_efd93a16("Tank 1P Status", 168, 315, -1, 0, 1)
   Button "Button_4" at 547,375 size 150x40; TextOff 'Disable Tank'; Authorization "Operate"
      on Press: function_b14e0dd5("504_Tank Grouping_DB2020_TANK ACTIV 2", 0)
   TextField "Text field_1" at 20,90 size 109x25; Text 'TIME LEFT:'
   GraphicView "Graphic view_1" at 20,46 size 245x32; Picture "Tank Manually Disabled"
   GraphicIOField "Graphic I/O field_1" at 20,46 size 245x32; PictureList "Tank Process Stage_II"
      Visibility <- "504_Tank Grouping_DB2020_GROUP of TANK 2"
      ProcessValue <- "2110_BTCS_CNTRL_DB_BTCS_STATE"
   Button "Button_2" at 4,5 size 45x35; TextOff 'Text'; PictureOff "Graphic_286"
      on Click: function_efd93a16("Tank 1P Status", 0, 0, -1, -1, 1)
   Button "Button_3" at 287,375 size 230x40; TextOff 'Text'; Authorization "Operate"; PictureList "Water Level Override"
      on Press: InvertBit("2062_Warning_Data_Water Level Override 1P")
      ProcessValue <- "2062_Warning_Data_Water Level Override 1P"
   Button "Button_5" at 27,375 size 230x40; TextOff 'Tank Shutdown Alarm'
      ProcessValue <- "2062_Warning_Data_Water Level Override 1P"
      Visibility <- "2062_Warning_Data_Alarm Tank P1"
   Button "Button_6" at 27,375 size 230x40; TextOff 'No/Low Water Level'; Authorization "Operate"
      ProcessValue <- "2062_Warning_Data_Water Level Override 1P"
      Visibility <- "LT422 1P  TANK LEVEL ALARM_ALARM L"
   IOField "I/O field_29" at 218,90 size 47x25; FormatPattern 99; Unit m
      ProcessValue <- "504_Tank Grouping_DB2020_Time Left Tank_Time Left m Tank 2"
   IOField "I/O field_8" at 173,90 size 42x25; FormatPattern 99; Unit h
      ProcessValue <- "504_Tank Grouping_DB2020_Time Left Tank_Time Left h Tank 2"
   IOField "I/O field_9" at 128,90 size 42x25; FormatPattern 99; Unit d
      ProcessValue <- "504_Tank Grouping_DB2020_Time Left Tank_Time Left d Tank 2"

PopupScreen "Tank 1S Status" 885x425
   TrendView "Trend view_1" at 280,7 size 600x360
   TextField "Text field_4" at 20,135 size 86x22; Text 'Pressure:'
   IOField "I/O field_1" at 175,130 size 90x25; FormatPattern s999.9; Unit  mBar
      ProcessValue <- "20_TANKS_IP_DATA_RIO_01_FIRST_TANK_TANKS_PRESS"
   TextField "Text field_5" at 20,169 size 113x22; Text 'Water Level:'
   IOField "I/O field_2" at 175,164 size 90x25; FormatPattern 999.9; Unit  %
      ProcessValue <- "20_TANKS_IP_DATA_RIO_01_THIRD_TANK_BWT_LEVEL"
   TextField "Text field_6" at 20,203 size 137x22; Text 'MBG Flow Rate:'
   IOField "I/O field_3" at 175,198 size 90x25; FormatPattern 999.9; Unit  m³/hr
      ProcessValue <- "20_TANKS_IP_DATA_RIO_01_THIRD_TANK_MBG_FLOW"
   TextField "Text field_7" at 20,237 size 135x22; Text 'USD Flow Rate:'
   IOField "I/O field_4" at 175,232 size 90x25; FormatPattern 999.9; Unit  m³/hr
      ProcessValue <- "20_TANKS_IP_DATA_RIO_01_THIRD_TANK_USD_FLOW"
   TextField "Text field_8" at 20,271 size 140x22; Text 'Water pH Level:'
   IOField "I/O field_5" at 175,266 size 90x25; FormatPattern 99.9
      ProcessValue <- "20_TANKS_IP_DATA_RIO_01_THIRD_TANK_BWT_PH"
   TextField "Text field_9" at 20,305 size 143x22; Text 'Water DO Level:'
   IOField "I/O field_6" at 175,300 size 90x25; FormatPattern 99.99; Unit  mg/l
      ProcessValue <- "20_TANKS_IP_DATA_RIO_01_THIRD_TANK_BWT_DO"
   TextField "Text field_10" at 20,339 size 174x22; Text 'Water Temperature:'
   IOField "I/O field_7" at 190,334 size 75x25; FormatPattern 999.9; Unit  °C
      ProcessValue <- "20_TANKS_IP_DATA_RIO_01_THIRD_TANK_BWT_TEMP"
   Button "Button_1" at 50,5 size 220x35; TextOff 'Starboard Tank 1 (1S)'
      on Release: function_efd93a16("Tank 1S Status", 168, 315, -1, 0, 1)
   Button "Button_4" at 548,375 size 150x40; TextOff 'Disable Tank'; Authorization "Operate"
      on Press: function_b14e0dd5("504_Tank Grouping_DB2020_TANK ACTIV 3", 0)
   TextField "Text field_1" at 20,90 size 109x25; Text 'TIME LEFT:'
   GraphicView "Graphic view_1" at 20,46 size 245x32; Picture "Tank Manually Disabled"
   GraphicIOField "Graphic I/O field_1" at 20,46 size 245x32; PictureList "Tank Process Stage_II"
      Visibility <- "504_Tank Grouping_DB2020_GROUP of TANK 3"
      ProcessValue <- "2110_BTCS_CNTRL_DB_BTCS_STATE"
   Button "Button_2" at 4,5 size 45x35; TextOff 'Text'; PictureOff "Graphic_286"
      on Click: function_efd93a16("Tank 1S Status", 0, 0, -1, -1, 1)
   Button "Button_3" at 287,375 size 230x40; TextOff 'Text'; Authorization "Operate"; PictureList "Water Level Override"
      on Press: InvertBit("2062_Warning_Data_Water Level Override 1S")
      ProcessValue <- "2062_Warning_Data_Water Level Override 1S"
   Button "Button_5" at 27,375 size 230x40; TextOff 'Tank Shutdown Alarm'
      Visibility <- "2062_Warning_Data_Alarm Tank S1"
   Button "Button_6" at 27,375 size 230x40; TextOff 'No/Low Water Level'; Authorization "Operate"
      Visibility <- "LT421 1S  TANK LEVEL ALARM_ALARM L"
   IOField "I/O field_29" at 218,90 size 47x25; FormatPattern 99; Unit m
      ProcessValue <- "504_Tank Grouping_DB2020_Time Left Tank_Time Left m Tank 3"
   IOField "I/O field_8" at 173,90 size 42x25; FormatPattern 99; Unit h
      ProcessValue <- "504_Tank Grouping_DB2020_Time Left Tank_Time Left h Tank 3"
   IOField "I/O field_9" at 128,90 size 42x25; FormatPattern 99; Unit d
      ProcessValue <- "504_Tank Grouping_DB2020_Time Left Tank_Time Left d Tank 3"

PopupScreen "Tank 2P Status" 885x425
   TrendView "Trend view_1" at 280,7 size 600x360
   TextField "Text field_4" at 20,135 size 86x22; Text 'Pressure:'
   IOField "I/O field_1" at 175,130 size 90x25; FormatPattern s999.9; Unit  mBar
      ProcessValue <- "20_TANKS_IP_DATA_RIO_02_FIRST_TANK_TANKS_PRESS"
   TextField "Text field_5" at 20,169 size 113x22; Text 'Water Level:'
   IOField "I/O field_2" at 175,164 size 90x25; FormatPattern 999.9; Unit  %
      ProcessValue <- "20_TANKS_IP_DATA_RIO_02_FIRST_TANK_BWT_LEVEL"
   TextField "Text field_6" at 20,203 size 137x22; Text 'MBG Flow Rate:'
   IOField "I/O field_3" at 175,198 size 90x25; FormatPattern 999.9; Unit  m³/hr
      ProcessValue <- "20_TANKS_IP_DATA_RIO_02_FIRST_TANK_MBG_FLOW"
   TextField "Text field_7" at 20,237 size 135x22; Text 'USD Flow Rate:'
   IOField "I/O field_4" at 175,232 size 90x25; FormatPattern 999.9; Unit  m³/hr
      ProcessValue <- "20_TANKS_IP_DATA_RIO_02_FIRST_TANK_USD_FLOW"
   TextField "Text field_8" at 20,271 size 140x22; Text 'Water pH Level:'
   IOField "I/O field_5" at 175,266 size 90x25; FormatPattern 99.9
      ProcessValue <- "20_TANKS_IP_DATA_RIO_02_FIRST_TANK_BWT_PH"
   TextField "Text field_9" at 20,305 size 143x22; Text 'Water DO Level:'
   IOField "I/O field_6" at 175,300 size 90x25; FormatPattern 99.99; Unit  mg/l
      ProcessValue <- "20_TANKS_IP_DATA_RIO_02_FIRST_TANK_BWT_DO"
   TextField "Text field_10" at 20,339 size 174x22; Text 'Water Temperature:'
   IOField "I/O field_7" at 190,334 size 75x25; FormatPattern 999.9; Unit  °C
      ProcessValue <- "20_TANKS_IP_DATA_RIO_02_FIRST_TANK_BWT_TEMP"
   Button "Button_4" at 545,375 size 150x40; TextOff 'Disable Tank'; Authorization "Operate"
      on Press: function_b14e0dd5("504_Tank Grouping_DB2020_TANK ACTIV 4", 0)
   Button "Button_1" at 51,5 size 219x35; TextOff 'Port Tank 2 (2P)'
      on Release: function_efd93a16("Tank 2P Status", 168, 315, -1, 0, 1)
   TextField "Text field_1" at 20,90 size 109x25; Text 'TIME LEFT:'
   GraphicView "Graphic view_1" at 20,46 size 245x32; Picture "Tank Manually Disabled"
   GraphicIOField "Graphic I/O field_1" at 20,46 size 245x32; PictureList "Tank Process Stage_II"
      Visibility <- "504_Tank Grouping_DB2020_GROUP of TANK 4"
      ProcessValue <- "2110_BTCS_CNTRL_DB_BTCS_STATE"
   Button "Button_2" at 4,5 size 45x35; TextOff 'Text'; PictureOff "Graphic_286"
      on Click: function_efd93a16("Tank 2P Status", 0, 0, -1, -1, 1)
   Button "Button_3" at 287,375 size 230x40; TextOff 'Text'; Authorization "Operate"; PictureList "Water Level Override"
      on Press: InvertBit("2062_Warning_Data_Water Level Override 2P")
      ProcessValue <- "2062_Warning_Data_Water Level Override 2P"
   Button "Button_5" at 27,375 size 230x40; TextOff 'Tank Shutdown Alarm'
      Visibility <- "2062_Warning_Data_Alarm Tank P2"
   Button "Button_6" at 27,375 size 230x40; TextOff 'No/Low Water Level'; Authorization "Operate"
      Visibility <- "FIT418_2P_ALM_ANALOG_DB_ALARM L"
   IOField "I/O field_29" at 218,90 size 47x25; FormatPattern 99; Unit m
      ProcessValue <- "504_Tank Grouping_DB2020_Time Left Tank_Time Left m Tank 4"
   IOField "I/O field_8" at 173,90 size 42x25; FormatPattern 99; Unit h
      ProcessValue <- "504_Tank Grouping_DB2020_Time Left Tank_Time Left h Tank 4"
   IOField "I/O field_9" at 128,90 size 42x25; FormatPattern 99; Unit d
      ProcessValue <- "504_Tank Grouping_DB2020_Time Left Tank_Time Left d Tank 4"

